                           ValveDemand := #GTT_IN.GTT_ValveDemands[1],
                           OpenTime := "1096_ADJUSTABLE_CONSTANTS".BWTInletValveOpen_Time,
                           CloseTime := "1096_ADJUSTABLE_CONSTANTS".BWTInletValveClose_Time,
                           ENO => #_w2);
   #DNC_FPT_GTT(EN := #_w2,   // "1604_DEMAND_AND_CHECK"
                DemandIn := #GTT_IN.GTT_ValveDemands[1],
                NO_Type := False,
                NC_Type := True,
                ValveMoveTime := #FPT_GTT_TimeSel,
                ValveOpenStatus := "20_TANKS_IP_DATA".RIO_01.FIRST_TANK.TANK_VENT_A_OPEN,
                ValveClsdStatus := "20_TANKS_IP_DATA".RIO_01.FIRST_TANK.TANK_VENT_A_CLSD,
                DemandOut => "40_TANKS_OP_DATA".RIO_01_VENT_A_FPT,
                DemandComplete => #GTT_OUT.GTT_DemandsCompleted[1],
                Alarm => #GTT_OUT.GTT_Alarms[1],
                ENO => #_w3);
   IF #_w3 THEN
       "1133_GTT_DETERMINE_EXCLUSIVITY"(TankID_InOperation := 1,
                               DemandComplete := #GTT_OUT.GTT_DemandsCompleted[1],
                               GTT_Exclusivity := #GTT_Exclusivity);
   END_IF;
   #DNC_FPT_GTT.Reset := NOT #_w1;
   #_w4 := (NOT #GTT_Exclusivity.Tank_Exclusivity AND #GTT_IN.GTT_Actuate[2] AND NOT #GTT_OUT.GTT_DemandsCompleted[2]) OR (#GTT_Exclusivity.TankID_InOperation = 2);
   #"1P_GTT_TimeSel" := "1135_VALVE_OPEN_CLOSE_TIME_SEL"(EN := #_w4,
                           ValveType := 0,
                           ValveDemand := #GTT_IN.GTT_ValveDemands[2],
                           OpenTime := "1096_ADJUSTABLE_CONSTANTS".BWTInletValveOpen_Time,
                           CloseTime := "1096_ADJUSTABLE_CONSTANTS".BWTInletValveClose_Time,
                           ENO => #_w5);
   #DNC_1P_GTT(EN := #_w5,   // "1604_DEMAND_AND_CHECK"
               DemandIn := #GTT_IN.GTT_ValveDemands[2],
               NO_Type := False,
               NC_Type := True,
               ValveMoveTime := #"1P_GTT_TimeSel",
               ValveOpenStatus := "20_TANKS_IP_DATA".RIO_01.SECOND_TANK.TANK_VENT_A_OPEN,
               ValveClsdStatus := "20_TANKS_IP_DATA".RIO_01.SECOND_TANK.TANK_VENT_A_CLSD,
               DemandOut => "40_TANKS_OP_DATA".RIO_01_VENT_A_1P,
               DemandComplete => #GTT_OUT.GTT_DemandsCompleted[2],
               Alarm => #GTT_OUT.GTT_Alarms[2],
               ENO => #_w6);
   IF #_w6 THEN
       "1133_GTT_DETERMINE_EXCLUSIVITY"(TankID_InOperation := 2,
                               DemandComplete := #GTT_OUT.GTT_DemandsCompleted[2],
                               GTT_Exclusivity := #GTT_Exclusivity);
   END_IF;
   #DNC_1P_GTT.Reset := NOT #_w4;
   #_w7 := (NOT #GTT_Exclusivity.Tank_Exclusivity AND #GTT_IN.GTT_Actuate[3] AND NOT #GTT_OUT.GTT_DemandsCompleted[3]) OR (#GTT_Exclusivity.TankID_InOperation = 3);
   #"1S_GTT_TimeSel" := "1135_VALVE_OPEN_CLOSE_TIME_SEL"(EN := #_w7,
                           ValveType := 0,
                           ValveDemand := #GTT_IN.GTT_ValveDemands[3],
                           OpenTime := "1096_ADJUSTABLE_CONSTANTS".BWTInletValveOpen_Time,
                           CloseTime := "1096_ADJUSTABLE_CONSTANTS".BWTInletValveClose_Time,
                           ENO => #_w8);
   #DNC_1S_GTT(EN := #_w8,   // "1604_DEMAND_AND_CHECK"
               DemandIn := #GTT_IN.GTT_ValveDemands[3],
               NO_Type := False,
               NC_Type := True,
               ValveMoveTime := #"1S_GTT_TimeSel",
               ValveOpenStatus := "20_TANKS_IP_DATA".RIO_01.THIRD_TANK.TANK_VENT_A_OPEN,
               ValveClsdStatus := "20_TANKS_IP_DATA".RIO_01.THIRD_TANK.TANK_VENT_A_CLSD,
               DemandOut => "40_TANKS_OP_DATA".RIO_01_VENT_A_1S,
               DemandComplete => #GTT_OUT.GTT_DemandsCompleted[3],
               Alarm => #GTT_OUT.GTT_Alarms[3],
               ENO => #_w9);
   IF #_w9 THEN
       "1133_GTT_DETERMINE_EXCLUSIVITY"(TankID_InOperation := 3,
                               DemandComplete := #GTT_OUT.GTT_DemandsCompleted[3],
                               GTT_Exclusivity := #GTT_Exclusivity);
   END_IF;
   #DNC_1S_GTT.Reset := NOT #_w7;
END_REGION

REGION Network 3: RIO02 2P, 2S GTT control
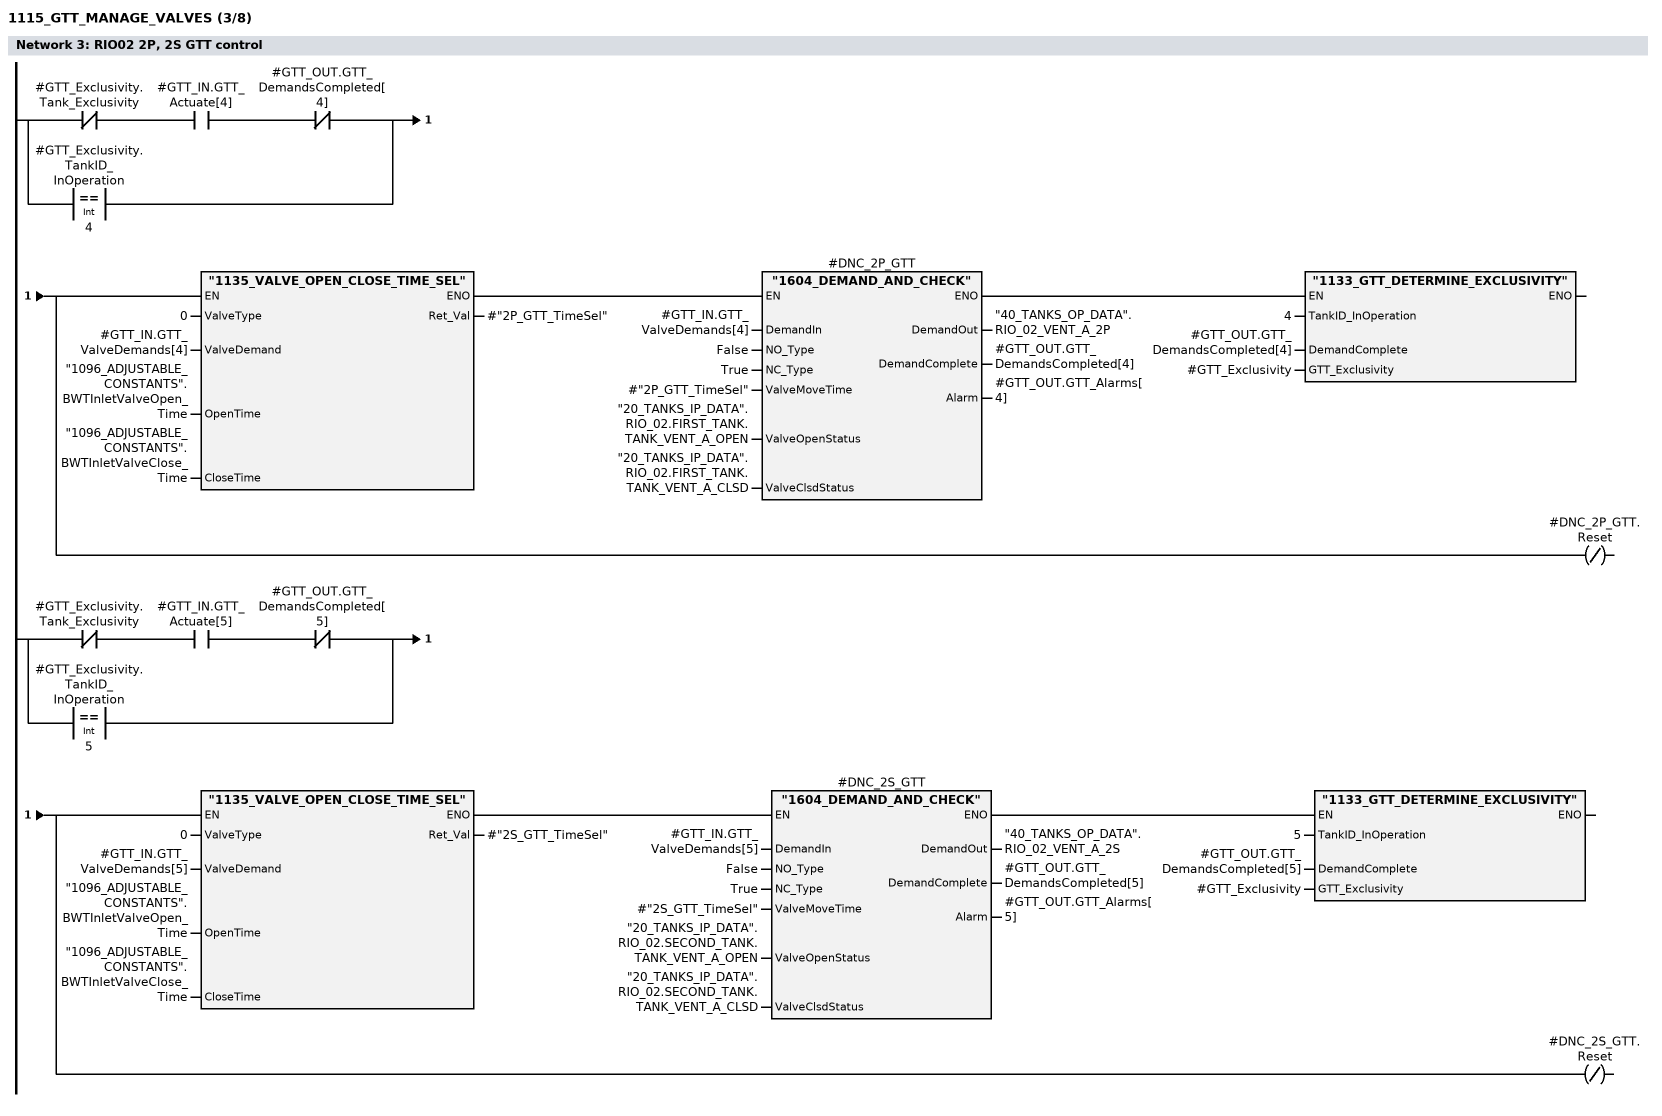
   RUNG wire#powerrail
      I_Contact( #GTT_Exclusivity.Tank_Exclusivity )
      Contact( #GTT_IN.GTT_Actuate[4] )
      I_Contact( #GTT_OUT.GTT_DemandsCompleted[4] )
      wire#w1
      "1135_VALVE_OPEN_CLOSE_TIME_SEL"(ValveType := 0, ValveDemand := #GTT_IN.GTT_ValveDemands[4], OpenTime := "1096_ADJUSTABLE_CONSTANTS".BWTInletValveOpen_Time, CloseTime := "1096_ADJUSTABLE_CONSTANTS".BWTInletValveClose_Time, Ret_Val => #"2P_GTT_TimeSel")
      #DNC_2P_GTT(DemandIn := #GTT_IN.GTT_ValveDemands[4], NO_Type := False, NC_Type := True, ValveMoveTime := #"2P_GTT_TimeSel", ValveOpenStatus := "20_TANKS_IP_DATA".RIO_02.FIRST_TANK.TANK_VENT_A_OPEN, ValveClsdStatus := "20_TANKS_IP_DATA".RIO_02.FIRST_TANK.TANK_VENT_A_CLSD, DemandOut => "40_TANKS_OP_DATA".RIO_02_VENT_A_2P, DemandComplete => #GTT_OUT.GTT_DemandsCompleted[4], Alarm => #GTT_OUT.GTT_Alarms[4])
      "1133_GTT_DETERMINE_EXCLUSIVITY"(TankID_InOperation := 4, DemandComplete := #GTT_OUT.GTT_DemandsCompleted[4], GTT_Exclusivity := #GTT_Exclusivity)
   END_RUNG
   RUNG wire#powerrail
      { S7_Templates := "SrcType := Int" } EQ_Contact(in1 := #GTT_Exclusivity.TankID_InOperation, in2 := 4)
   END_RUNG wire#w1
   RUNG wire#w1
      I_Coil( #DNC_2P_GTT.Reset )
   END_RUNG
   RUNG wire#powerrail
      I_Contact( #GTT_Exclusivity.Tank_Exclusivity )
      Contact( #GTT_IN.GTT_Actuate[5] )
      I_Contact( #GTT_OUT.GTT_DemandsCompleted[5] )
      wire#w2
      "1135_VALVE_OPEN_CLOSE_TIME_SEL"(ValveType := 0, ValveDemand := #GTT_IN.GTT_ValveDemands[5], OpenTime := "1096_ADJUSTABLE_CONSTANTS".BWTInletValveOpen_Time, CloseTime := "1096_ADJUSTABLE_CONSTANTS".BWTInletValveClose_Time, Ret_Val => #"2S_GTT_TimeSel")
      #DNC_2S_GTT(DemandIn := #GTT_IN.GTT_ValveDemands[5], NO_Type := False, NC_Type := True, ValveMoveTime := #"2S_GTT_TimeSel", ValveOpenStatus := "20_TANKS_IP_DATA".RIO_02.SECOND_TANK.TANK_VENT_A_OPEN, ValveClsdStatus := "20_TANKS_IP_DATA".RIO_02.SECOND_TANK.TANK_VENT_A_CLSD, DemandOut => "40_TANKS_OP_DATA".RIO_02_VENT_A_2S, DemandComplete => #GTT_OUT.GTT_DemandsCompleted[5], Alarm => #GTT_OUT.GTT_Alarms[5])
      "1133_GTT_DETERMINE_EXCLUSIVITY"(TankID_InOperation := 5, DemandComplete := #GTT_OUT.GTT_DemandsCompleted[5], GTT_Exclusivity := #GTT_Exclusivity)
   END_RUNG
   RUNG wire#powerrail
      { S7_Templates := "SrcType := Int" } EQ_Contact(in1 := #GTT_Exclusivity.TankID_InOperation, in2 := 5)
   END_RUNG wire#w2
   RUNG wire#w2
      I_Coil( #DNC_2S_GTT.Reset )
   END_RUNG
   // the same network as SCL:
   #_w1 := (NOT #GTT_Exclusivity.Tank_Exclusivity AND #GTT_IN.GTT_Actuate[4] AND NOT #GTT_OUT.GTT_DemandsCompleted[4]) OR (#GTT_Exclusivity.TankID_InOperation = 4);
   #"2P_GTT_TimeSel" := "1135_VALVE_OPEN_CLOSE_TIME_SEL"(EN := #_w1,
                           ValveType := 0,
                           ValveDemand := #GTT_IN.GTT_ValveDemands[4],
                           OpenTime := "1096_ADJUSTABLE_CONSTANTS".BWTInletValveOpen_Time,
                           CloseTime := "1096_ADJUSTABLE_CONSTANTS".BWTInletValveClose_Time,
                           ENO => #_w2);
   #DNC_2P_GTT(EN := #_w2,   // "1604_DEMAND_AND_CHECK"
               DemandIn := #GTT_IN.GTT_ValveDemands[4],
               NO_Type := False,
               NC_Type := True,
               ValveMoveTime := #"2P_GTT_TimeSel",
               ValveOpenStatus := "20_TANKS_IP_DATA".RIO_02.FIRST_TANK.TANK_VENT_A_OPEN,
               ValveClsdStatus := "20_TANKS_IP_DATA".RIO_02.FIRST_TANK.TANK_VENT_A_CLSD,
               DemandOut => "40_TANKS_OP_DATA".RIO_02_VENT_A_2P,
               DemandComplete => #GTT_OUT.GTT_DemandsCompleted[4],
               Alarm => #GTT_OUT.GTT_Alarms[4],
               ENO => #_w3);
   IF #_w3 THEN
       "1133_GTT_DETERMINE_EXCLUSIVITY"(TankID_InOperation := 4,
                               DemandComplete := #GTT_OUT.GTT_DemandsCompleted[4],
                               GTT_Exclusivity := #GTT_Exclusivity);
   END_IF;
   #DNC_2P_GTT.Reset := NOT #_w1;
   #_w4 := (NOT #GTT_Exclusivity.Tank_Exclusivity AND #GTT_IN.GTT_Actuate[5] AND NOT #GTT_OUT.GTT_DemandsCompleted[5]) OR (#GTT_Exclusivity.TankID_InOperation = 5);
   #"2S_GTT_TimeSel" := "1135_VALVE_OPEN_CLOSE_TIME_SEL"(EN := #_w4,
                           ValveType := 0,
                           ValveDemand := #GTT_IN.GTT_ValveDemands[5],
                           OpenTime := "1096_ADJUSTABLE_CONSTANTS".BWTInletValveOpen_Time,
                           CloseTime := "1096_ADJUSTABLE_CONSTANTS".BWTInletValveClose_Time,
                           ENO => #_w5);
   #DNC_2S_GTT(EN := #_w5,   // "1604_DEMAND_AND_CHECK"
               DemandIn := #GTT_IN.GTT_ValveDemands[5],
               NO_Type := False,
               NC_Type := True,
               ValveMoveTime := #"2S_GTT_TimeSel",
               ValveOpenStatus := "20_TANKS_IP_DATA".RIO_02.SECOND_TANK.TANK_VENT_A_OPEN,
               ValveClsdStatus := "20_TANKS_IP_DATA".RIO_02.SECOND_TANK.TANK_VENT_A_CLSD,
               DemandOut => "40_TANKS_OP_DATA".RIO_02_VENT_A_2S,
               DemandComplete => #GTT_OUT.GTT_DemandsCompleted[5],
               Alarm => #GTT_OUT.GTT_Alarms[5],
               ENO => #_w6);
   IF #_w6 THEN
       "1133_GTT_DETERMINE_EXCLUSIVITY"(TankID_InOperation := 5,
                               DemandComplete := #GTT_OUT.GTT_DemandsCompleted[5],
                               GTT_Exclusivity := #GTT_Exclusivity);
   END_IF;
   #DNC_2S_GTT.Reset := NOT #_w4;
END_REGION

REGION Network 4: RIO02 3P, 3S GTT control
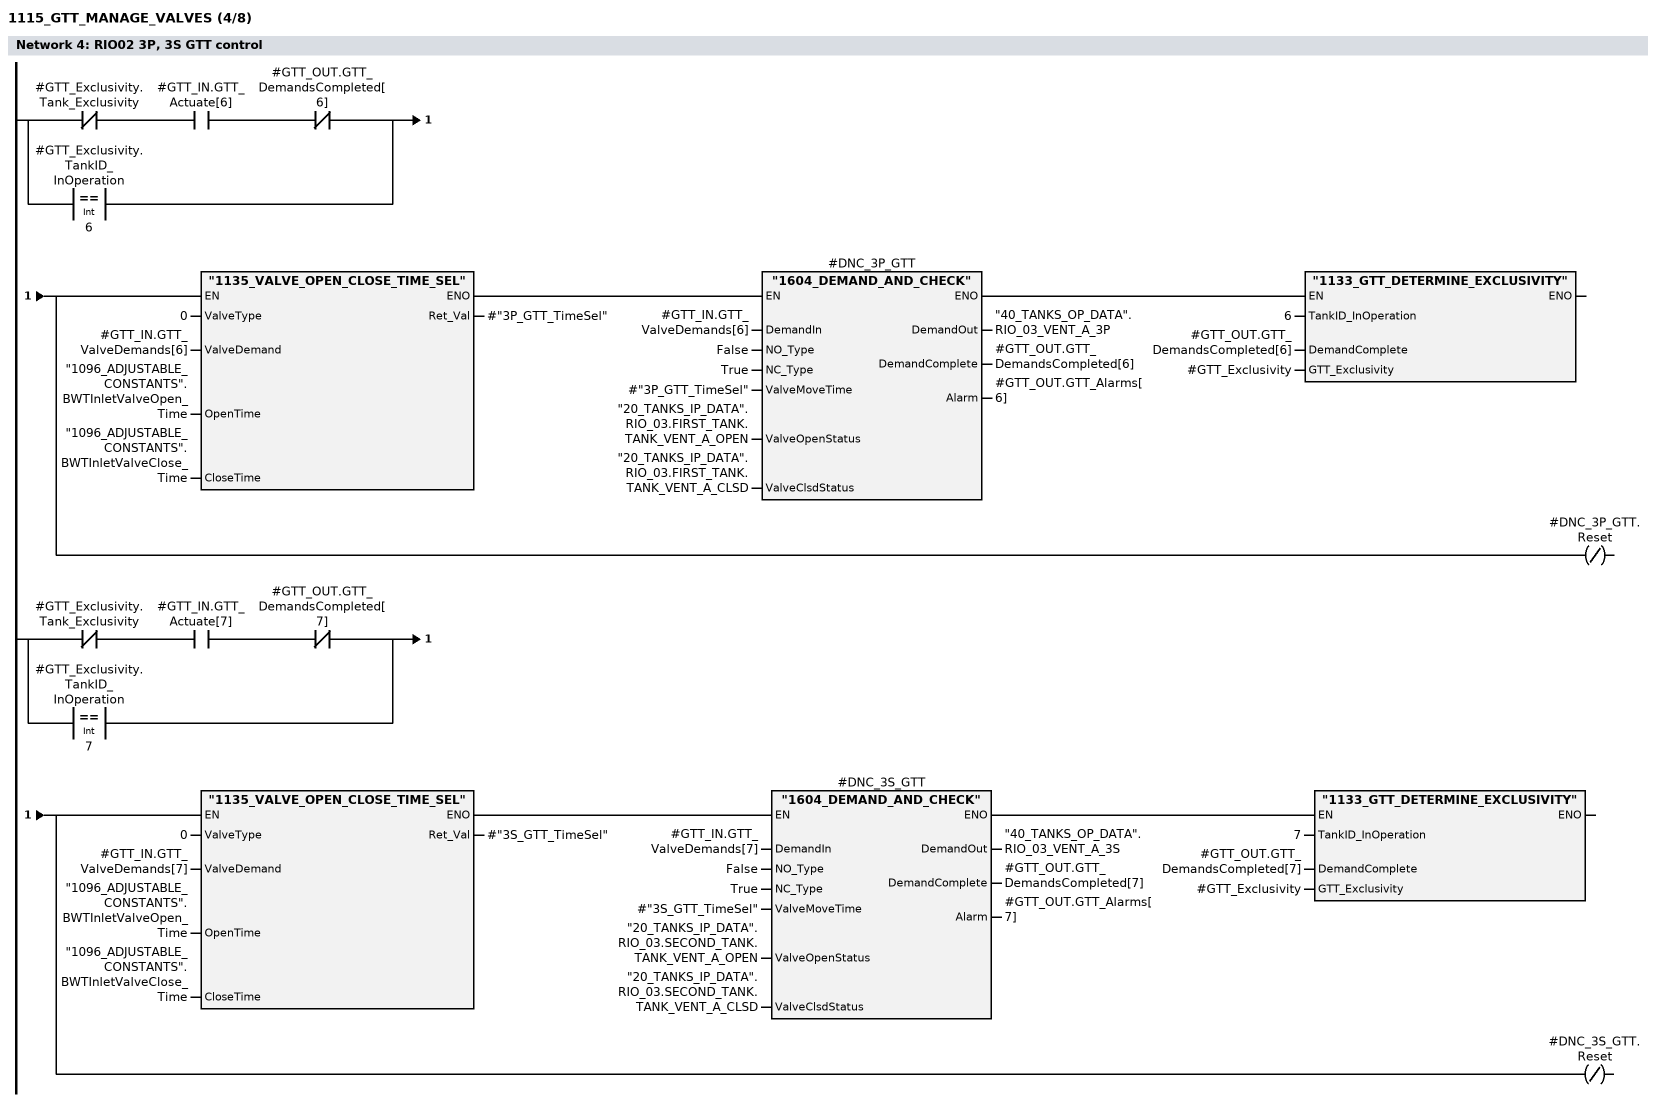
   RUNG wire#powerrail
      I_Contact( #GTT_Exclusivity.Tank_Exclusivity )
      Contact( #GTT_IN.GTT_Actuate[6] )
      I_Contact( #GTT_OUT.GTT_DemandsCompleted[6] )
      wire#w1
      "1135_VALVE_OPEN_CLOSE_TIME_SEL"(ValveType := 0, ValveDemand := #GTT_IN.GTT_ValveDemands[6], OpenTime := "1096_ADJUSTABLE_CONSTANTS".BWTInletValveOpen_Time, CloseTime := "1096_ADJUSTABLE_CONSTANTS".BWTInletValveClose_Time, Ret_Val => #"3P_GTT_TimeSel")
      #DNC_3P_GTT(DemandIn := #GTT_IN.GTT_ValveDemands[6], NO_Type := False, NC_Type := True, ValveMoveTime := #"3P_GTT_TimeSel", ValveOpenStatus := "20_TANKS_IP_DATA".RIO_03.FIRST_TANK.TANK_VENT_A_OPEN, ValveClsdStatus := "20_TANKS_IP_DATA".RIO_03.FIRST_TANK.TANK_VENT_A_CLSD, DemandOut => "40_TANKS_OP_DATA".RIO_03_VENT_A_3P, DemandComplete => #GTT_OUT.GTT_DemandsCompleted[6], Alarm => #GTT_OUT.GTT_Alarms[6])
      "1133_GTT_DETERMINE_EXCLUSIVITY"(TankID_InOperation := 6, DemandComplete := #GTT_OUT.GTT_DemandsCompleted[6], GTT_Exclusivity := #GTT_Exclusivity)
   END_RUNG
   RUNG wire#powerrail
      { S7_Templates := "SrcType := Int" } EQ_Contact(in1 := #GTT_Exclusivity.TankID_InOperation, in2 := 6)
   END_RUNG wire#w1
   RUNG wire#w1
      I_Coil( #DNC_3P_GTT.Reset )
   END_RUNG
   RUNG wire#powerrail
      I_Contact( #GTT_Exclusivity.Tank_Exclusivity )
      Contact( #GTT_IN.GTT_Actuate[7] )
      I_Contact( #GTT_OUT.GTT_DemandsCompleted[7] )
      wire#w2
      "1135_VALVE_OPEN_CLOSE_TIME_SEL"(ValveType := 0, ValveDemand := #GTT_IN.GTT_ValveDemands[7], OpenTime := "1096_ADJUSTABLE_CONSTANTS".BWTInletValveOpen_Time, CloseTime := "1096_ADJUSTABLE_CONSTANTS".BWTInletValveClose_Time, Ret_Val => #"3S_GTT_TimeSel")
      #DNC_3S_GTT(DemandIn := #GTT_IN.GTT_ValveDemands[7], NO_Type := False, NC_Type := True, ValveMoveTime := #"3S_GTT_TimeSel", ValveOpenStatus := "20_TANKS_IP_DATA".RIO_03.SECOND_TANK.TANK_VENT_A_OPEN, ValveClsdStatus := "20_TANKS_IP_DATA".RIO_03.SECOND_TANK.TANK_VENT_A_CLSD, DemandOut => "40_TANKS_OP_DATA".RIO_03_VENT_A_3S, DemandComplete => #GTT_OUT.GTT_DemandsCompleted[7], Alarm => #GTT_OUT.GTT_Alarms[7])
      "1133_GTT_DETERMINE_EXCLUSIVITY"(TankID_InOperation := 7, DemandComplete := #GTT_OUT.GTT_DemandsCompleted[7], GTT_Exclusivity := #GTT_Exclusivity)
   END_RUNG
   RUNG wire#powerrail
      { S7_Templates := "SrcType := Int" } EQ_Contact(in1 := #GTT_Exclusivity.TankID_InOperation, in2 := 7)
   END_RUNG wire#w2
   RUNG wire#w2
      I_Coil( #DNC_3S_GTT.Reset )
   END_RUNG
   // the same network as SCL:
   #_w1 := (NOT #GTT_Exclusivity.Tank_Exclusivity AND #GTT_IN.GTT_Actuate[6] AND NOT #GTT_OUT.GTT_DemandsCompleted[6]) OR (#GTT_Exclusivity.TankID_InOperation = 6);
   #"3P_GTT_TimeSel" := "1135_VALVE_OPEN_CLOSE_TIME_SEL"(EN := #_w1,
                           ValveType := 0,
                           ValveDemand := #GTT_IN.GTT_ValveDemands[6],
                           OpenTime := "1096_ADJUSTABLE_CONSTANTS".BWTInletValveOpen_Time,
                           CloseTime := "1096_ADJUSTABLE_CONSTANTS".BWTInletValveClose_Time,
                           ENO => #_w2);
   #DNC_3P_GTT(EN := #_w2,   // "1604_DEMAND_AND_CHECK"
               DemandIn := #GTT_IN.GTT_ValveDemands[6],
               NO_Type := False,
               NC_Type := True,
               ValveMoveTime := #"3P_GTT_TimeSel",
               ValveOpenStatus := "20_TANKS_IP_DATA".RIO_03.FIRST_TANK.TANK_VENT_A_OPEN,
               ValveClsdStatus := "20_TANKS_IP_DATA".RIO_03.FIRST_TANK.TANK_VENT_A_CLSD,
               DemandOut => "40_TANKS_OP_DATA".RIO_03_VENT_A_3P,
               DemandComplete => #GTT_OUT.GTT_DemandsCompleted[6],
               Alarm => #GTT_OUT.GTT_Alarms[6],
               ENO => #_w3);
   IF #_w3 THEN
       "1133_GTT_DETERMINE_EXCLUSIVITY"(TankID_InOperation := 6,
                               DemandComplete := #GTT_OUT.GTT_DemandsCompleted[6],
                               GTT_Exclusivity := #GTT_Exclusivity);
   END_IF;
   #DNC_3P_GTT.Reset := NOT #_w1;
   #_w4 := (NOT #GTT_Exclusivity.Tank_Exclusivity AND #GTT_IN.GTT_Actuate[7] AND NOT #GTT_OUT.GTT_DemandsCompleted[7]) OR (#GTT_Exclusivity.TankID_InOperation = 7);
   #"3S_GTT_TimeSel" := "1135_VALVE_OPEN_CLOSE_TIME_SEL"(EN := #_w4,
                           ValveType := 0,
                           ValveDemand := #GTT_IN.GTT_ValveDemands[7],
                           OpenTime := "1096_ADJUSTABLE_CONSTANTS".BWTInletValveOpen_Time,
                           CloseTime := "1096_ADJUSTABLE_CONSTANTS".BWTInletValveClose_Time,
                           ENO => #_w5);
   #DNC_3S_GTT(EN := #_w5,   // "1604_DEMAND_AND_CHECK"
               DemandIn := #GTT_IN.GTT_ValveDemands[7],
               NO_Type := False,
               NC_Type := True,
               ValveMoveTime := #"3S_GTT_TimeSel",
               ValveOpenStatus := "20_TANKS_IP_DATA".RIO_03.SECOND_TANK.TANK_VENT_A_OPEN,
               ValveClsdStatus := "20_TANKS_IP_DATA".RIO_03.SECOND_TANK.TANK_VENT_A_CLSD,
               DemandOut => "40_TANKS_OP_DATA".RIO_03_VENT_A_3S,
               DemandComplete => #GTT_OUT.GTT_DemandsCompleted[7],
               Alarm => #GTT_OUT.GTT_Alarms[7],
               ENO => #_w6);
   IF #_w6 THEN
       "1133_GTT_DETERMINE_EXCLUSIVITY"(TankID_InOperation := 7,
                               DemandComplete := #GTT_OUT.GTT_DemandsCompleted[7],
                               GTT_Exclusivity := #GTT_Exclusivity);
   END_IF;
   #DNC_3S_GTT.Reset := NOT #_w4;
END_REGION

REGION Network 5: RIO02 4P, 4S GTT control
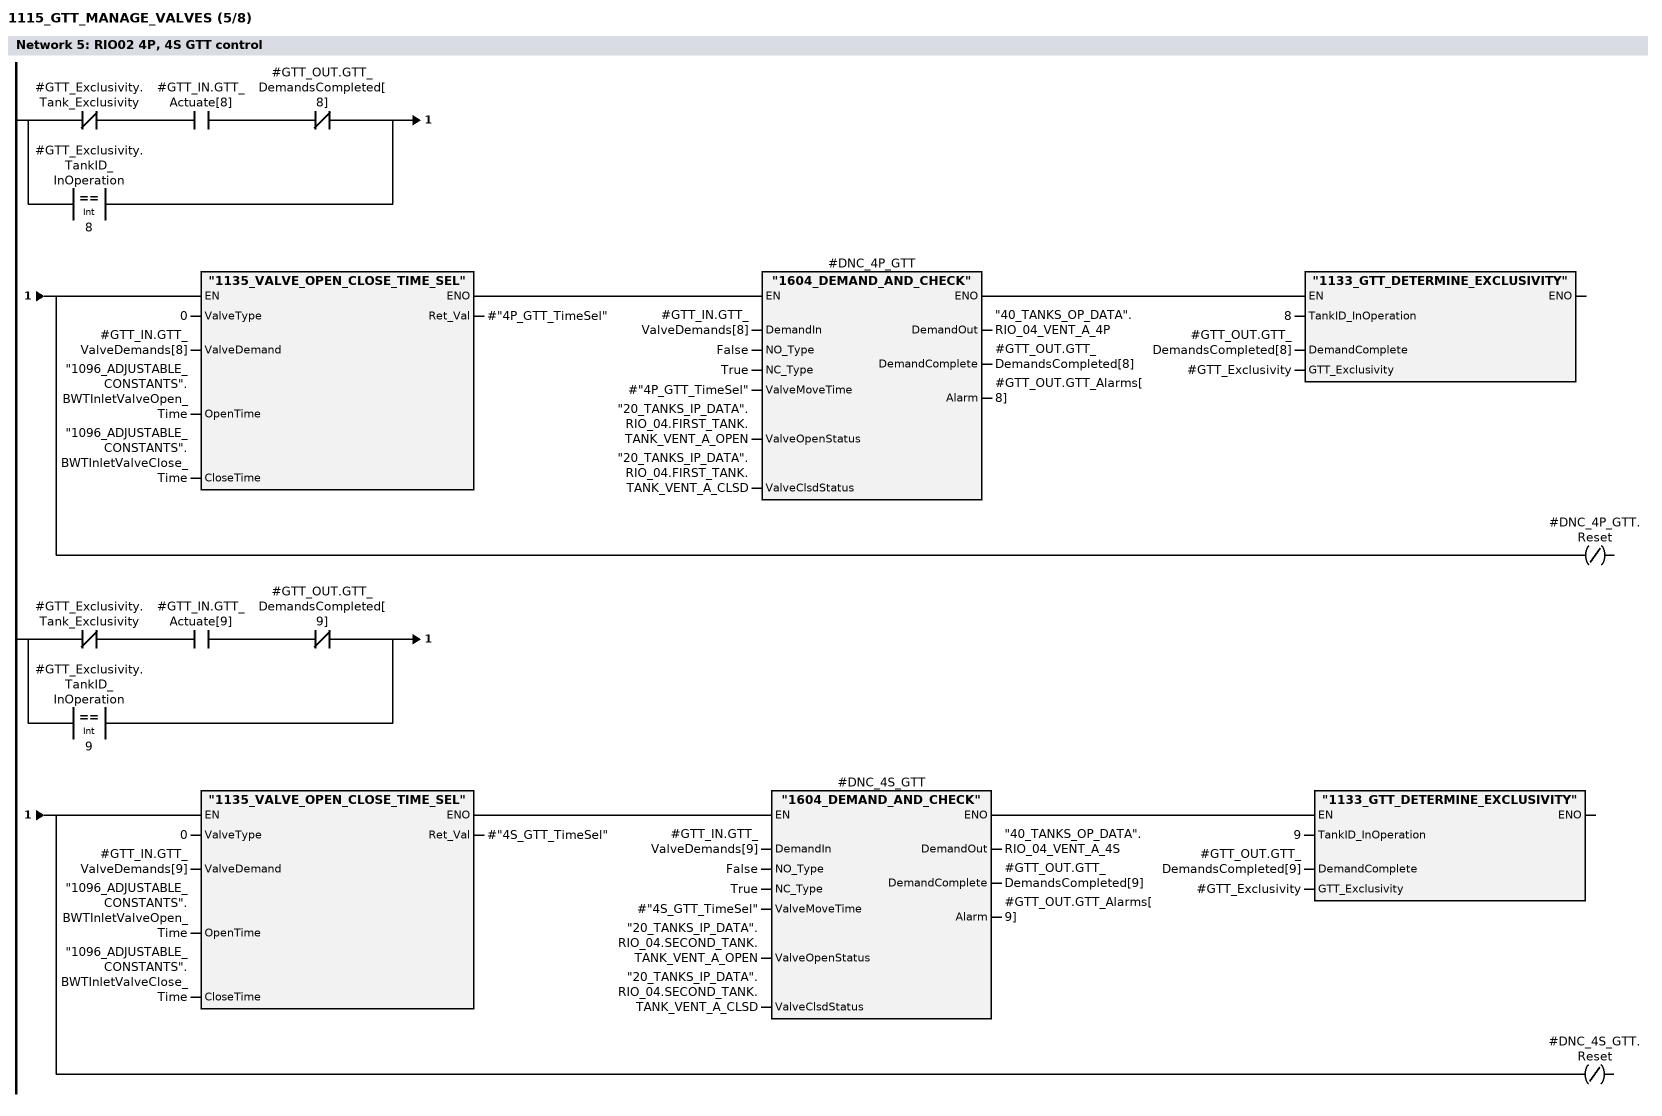
   RUNG wire#powerrail
      I_Contact( #GTT_Exclusivity.Tank_Exclusivity )
      Contact( #GTT_IN.GTT_Actuate[8] )
      I_Contact( #GTT_OUT.GTT_DemandsCompleted[8] )
      wire#w1
      "1135_VALVE_OPEN_CLOSE_TIME_SEL"(ValveType := 0, ValveDemand := #GTT_IN.GTT_ValveDemands[8], OpenTime := "1096_ADJUSTABLE_CONSTANTS".BWTInletValveOpen_Time, CloseTime := "1096_ADJUSTABLE_CONSTANTS".BWTInletValveClose_Time, Ret_Val => #"4P_GTT_TimeSel")
      #DNC_4P_GTT(DemandIn := #GTT_IN.GTT_ValveDemands[8], NO_Type := False, NC_Type := True, ValveMoveTime := #"4P_GTT_TimeSel", ValveOpenStatus := "20_TANKS_IP_DATA".RIO_04.FIRST_TANK.TANK_VENT_A_OPEN, ValveClsdStatus := "20_TANKS_IP_DATA".RIO_04.FIRST_TANK.TANK_VENT_A_CLSD, DemandOut => "40_TANKS_OP_DATA".RIO_04_VENT_A_4P, DemandComplete => #GTT_OUT.GTT_DemandsCompleted[8], Alarm => #GTT_OUT.GTT_Alarms[8])
      "1133_GTT_DETERMINE_EXCLUSIVITY"(TankID_InOperation := 8, DemandComplete := #GTT_OUT.GTT_DemandsCompleted[8], GTT_Exclusivity := #GTT_Exclusivity)
   END_RUNG
   RUNG wire#powerrail
      { S7_Templates := "SrcType := Int" } EQ_Contact(in1 := #GTT_Exclusivity.TankID_InOperation, in2 := 8)
   END_RUNG wire#w1
   RUNG wire#w1
      I_Coil( #DNC_4P_GTT.Reset )
   END_RUNG
   RUNG wire#powerrail
      I_Contact( #GTT_Exclusivity.Tank_Exclusivity )
      Contact( #GTT_IN.GTT_Actuate[9] )
      I_Contact( #GTT_OUT.GTT_DemandsCompleted[9] )
      wire#w2
      "1135_VALVE_OPEN_CLOSE_TIME_SEL"(ValveType := 0, ValveDemand := #GTT_IN.GTT_ValveDemands[9], OpenTime := "1096_ADJUSTABLE_CONSTANTS".BWTInletValveOpen_Time, CloseTime := "1096_ADJUSTABLE_CONSTANTS".BWTInletValveClose_Time, Ret_Val => #"4S_GTT_TimeSel")
      #DNC_4S_GTT(DemandIn := #GTT_IN.GTT_ValveDemands[9], NO_Type := False, NC_Type := True, ValveMoveTime := #"4S_GTT_TimeSel", ValveOpenStatus := "20_TANKS_IP_DATA".RIO_04.SECOND_TANK.TANK_VENT_A_OPEN, ValveClsdStatus := "20_TANKS_IP_DATA".RIO_04.SECOND_TANK.TANK_VENT_A_CLSD, DemandOut => "40_TANKS_OP_DATA".RIO_04_VENT_A_4S, DemandComplete => #GTT_OUT.GTT_DemandsCompleted[9], Alarm => #GTT_OUT.GTT_Alarms[9])
      "1133_GTT_DETERMINE_EXCLUSIVITY"(TankID_InOperation := 9, DemandComplete := #GTT_OUT.GTT_DemandsCompleted[9], GTT_Exclusivity := #GTT_Exclusivity)
   END_RUNG
   RUNG wire#powerrail
      { S7_Templates := "SrcType := Int" } EQ_Contact(in1 := #GTT_Exclusivity.TankID_InOperation, in2 := 9)
   END_RUNG wire#w2
   RUNG wire#w2
      I_Coil( #DNC_4S_GTT.Reset )
   END_RUNG
   // the same network as SCL:
   #_w1 := (NOT #GTT_Exclusivity.Tank_Exclusivity AND #GTT_IN.GTT_Actuate[8] AND NOT #GTT_OUT.GTT_DemandsCompleted[8]) OR (#GTT_Exclusivity.TankID_InOperation = 8);
   #"4P_GTT_TimeSel" := "1135_VALVE_OPEN_CLOSE_TIME_SEL"(EN := #_w1,
                           ValveType := 0,
                           ValveDemand := #GTT_IN.GTT_ValveDemands[8],
                           OpenTime := "1096_ADJUSTABLE_CONSTANTS".BWTInletValveOpen_Time,
                           CloseTime := "1096_ADJUSTABLE_CONSTANTS".BWTInletValveClose_Time,
                           ENO => #_w2);
   #DNC_4P_GTT(EN := #_w2,   // "1604_DEMAND_AND_CHECK"
               DemandIn := #GTT_IN.GTT_ValveDemands[8],
               NO_Type := False,
               NC_Type := True,
               ValveMoveTime := #"4P_GTT_TimeSel",
               ValveOpenStatus := "20_TANKS_IP_DATA".RIO_04.FIRST_TANK.TANK_VENT_A_OPEN,
               ValveClsdStatus := "20_TANKS_IP_DATA".RIO_04.FIRST_TANK.TANK_VENT_A_CLSD,
               DemandOut => "40_TANKS_OP_DATA".RIO_04_VENT_A_4P,
               DemandComplete => #GTT_OUT.GTT_DemandsCompleted[8],
               Alarm => #GTT_OUT.GTT_Alarms[8],
               ENO => #_w3);
   IF #_w3 THEN
       "1133_GTT_DETERMINE_EXCLUSIVITY"(TankID_InOperation := 8,
                               DemandComplete := #GTT_OUT.GTT_DemandsCompleted[8],
                               GTT_Exclusivity := #GTT_Exclusivity);
   END_IF;
   #DNC_4P_GTT.Reset := NOT #_w1;
   #_w4 := (NOT #GTT_Exclusivity.Tank_Exclusivity AND #GTT_IN.GTT_Actuate[9] AND NOT #GTT_OUT.GTT_DemandsCompleted[9]) OR (#GTT_Exclusivity.TankID_InOperation = 9);
   #"4S_GTT_TimeSel" := "1135_VALVE_OPEN_CLOSE_TIME_SEL"(EN := #_w4,
                           ValveType := 0,
                           ValveDemand := #GTT_IN.GTT_ValveDemands[9],
                           OpenTime := "1096_ADJUSTABLE_CONSTANTS".BWTInletValveOpen_Time,
                           CloseTime := "1096_ADJUSTABLE_CONSTANTS".BWTInletValveClose_Time,
                           ENO => #_w5);
   #DNC_4S_GTT(EN := #_w5,   // "1604_DEMAND_AND_CHECK"
               DemandIn := #GTT_IN.GTT_ValveDemands[9],
               NO_Type := False,
               NC_Type := True,
               ValveMoveTime := #"4S_GTT_TimeSel",
               ValveOpenStatus := "20_TANKS_IP_DATA".RIO_04.SECOND_TANK.TANK_VENT_A_OPEN,
               ValveClsdStatus := "20_TANKS_IP_DATA".RIO_04.SECOND_TANK.TANK_VENT_A_CLSD,
               DemandOut => "40_TANKS_OP_DATA".RIO_04_VENT_A_4S,
               DemandComplete => #GTT_OUT.GTT_DemandsCompleted[9],
               Alarm => #GTT_OUT.GTT_Alarms[9],
               ENO => #_w6);
   IF #_w6 THEN
       "1133_GTT_DETERMINE_EXCLUSIVITY"(TankID_InOperation := 9,
                               DemandComplete := #GTT_OUT.GTT_DemandsCompleted[9],
                               GTT_Exclusivity := #GTT_Exclusivity);
   END_IF;
   #DNC_4S_GTT.Reset := NOT #_w4;
END_REGION

REGION Network 6: RIO02 5P, 5S GTT control
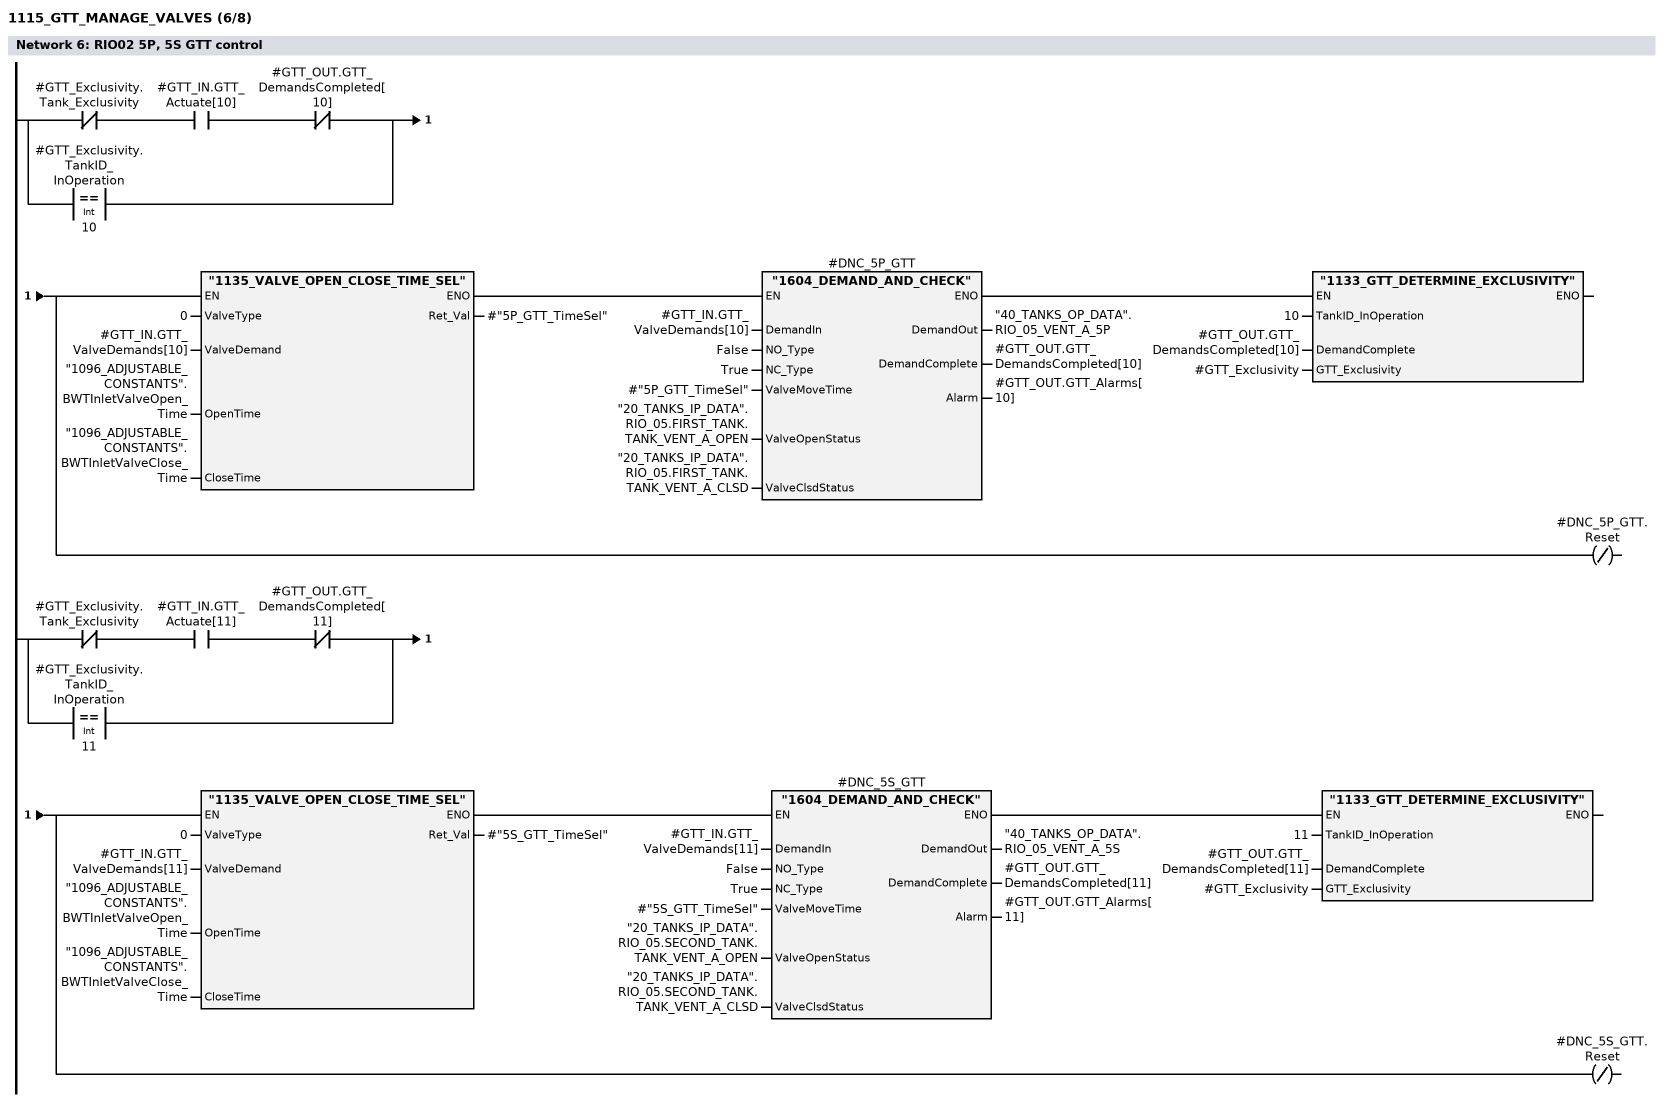
   RUNG wire#powerrail
      I_Contact( #GTT_Exclusivity.Tank_Exclusivity )
      Contact( #GTT_IN.GTT_Actuate[10] )
      I_Contact( #GTT_OUT.GTT_DemandsCompleted[10] )
      wire#w1
      "1135_VALVE_OPEN_CLOSE_TIME_SEL"(ValveType := 0, ValveDemand := #GTT_IN.GTT_ValveDemands[10], OpenTime := "1096_ADJUSTABLE_CONSTANTS".BWTInletValveOpen_Time, CloseTime := "1096_ADJUSTABLE_CONSTANTS".BWTInletValveClose_Time, Ret_Val => #"5P_GTT_TimeSel")
      #DNC_5P_GTT(DemandIn := #GTT_IN.GTT_ValveDemands[10], NO_Type := False, NC_Type := True, ValveMoveTime := #"5P_GTT_TimeSel", ValveOpenStatus := "20_TANKS_IP_DATA".RIO_05.FIRST_TANK.TANK_VENT_A_OPEN, ValveClsdStatus := "20_TANKS_IP_DATA".RIO_05.FIRST_TANK.TANK_VENT_A_CLSD, DemandOut => "40_TANKS_OP_DATA".RIO_05_VENT_A_5P, DemandComplete => #GTT_OUT.GTT_DemandsCompleted[10], Alarm => #GTT_OUT.GTT_Alarms[10])
      "1133_GTT_DETERMINE_EXCLUSIVITY"(TankID_InOperation := 10, DemandComplete := #GTT_OUT.GTT_DemandsCompleted[10], GTT_Exclusivity := #GTT_Exclusivity)
   END_RUNG
   RUNG wire#powerrail
      { S7_Templates := "SrcType := Int" } EQ_Contact(in1 := #GTT_Exclusivity.TankID_InOperation, in2 := 10)
   END_RUNG wire#w1
   RUNG wire#w1
      I_Coil( #DNC_5P_GTT.Reset )
   END_RUNG
   RUNG wire#powerrail
      I_Contact( #GTT_Exclusivity.Tank_Exclusivity )
      Contact( #GTT_IN.GTT_Actuate[11] )
      I_Contact( #GTT_OUT.GTT_DemandsCompleted[11] )
      wire#w2
      "1135_VALVE_OPEN_CLOSE_TIME_SEL"(ValveType := 0, ValveDemand := #GTT_IN.GTT_ValveDemands[11], OpenTime := "1096_ADJUSTABLE_CONSTANTS".BWTInletValveOpen_Time, CloseTime := "1096_ADJUSTABLE_CONSTANTS".BWTInletValveClose_Time, Ret_Val => #"5S_GTT_TimeSel")
      #DNC_5S_GTT(DemandIn := #GTT_IN.GTT_ValveDemands[11], NO_Type := False, NC_Type := True, ValveMoveTime := #"5S_GTT_TimeSel", ValveOpenStatus := "20_TANKS_IP_DATA".RIO_05.SECOND_TANK.TANK_VENT_A_OPEN, ValveClsdStatus := "20_TANKS_IP_DATA".RIO_05.SECOND_TANK.TANK_VENT_A_CLSD, DemandOut => "40_TANKS_OP_DATA".RIO_05_VENT_A_5S, DemandComplete => #GTT_OUT.GTT_DemandsCompleted[11], Alarm => #GTT_OUT.GTT_Alarms[11])